                   REGION "TEST STRING TOO LONG"
                       IF LEN(#lengthTest) > #maxLength THEN
                           #_lineBox[#pLineBox] := "Trim"(#_lineBox[#pLineBox]);
                           #_lineBox[#pLineBox] := "Trim"(#_lineBox[#pLineBox]);
                           #pLineBox := #pLineBox + 1;
                           #_lineBox[#pLineBox] := #stringBox[#pString];
                       END_IF;
                   END_REGION

               END_IF;
           END_REGION

       END_FOR;
   END_REGION

   REGION "RETURN"
       #lineBox := #_lineBox;
   END_REGION
END_FUNCTION

FUNCTION "WString.Word_Wrap_Depricated.Concat_Lines" : WString   // FC75, SCL
{ S7_Optimized_Access := 'TRUE' }
VERSION : 0.1
   VAR_INPUT
      lineBox : Array[0..#limitLines] of WString["LONG_STRING_LENGTH"];
   END_VAR
   VAR_TEMP
      pLine : Int;
      ret : WString;
   END_VAR
   VAR CONSTANT
      space : WString := WSTRING#' ';
      blank : WString;
      lineBreak : WString := WSTRING#'$L';
      limitString : Int := 49;
      limitLines : Int := 9;
   END_VAR
BEGIN
   REGION "FOR EACH LINE"
       FOR #pLine := 0 TO #limitLines DO

           REGION "ON END OF LINE LIST"
               IF #lineBox[#pLine] = #space OR #lineBox[#pLine] = #blank THEN
                   EXIT;
               END_IF;
           END_REGION

           REGION "ON FIRST ELEMENT IN LINE LIST"
               IF #pLine = 0 THEN
                   #ret := #lineBox[#pLine];
               END_IF;
           END_REGION

           REGION "CONSTRUCT OUTPUT"
               IF #pLine >= 1 THEN

                   REGION "NO OP ON LINE BREAK CHARACTER"
                       IF #lineBox[#pLine] = #lineBreak THEN
                           ;// no action required
                       END_IF;
                   END_REGION

                   REGION "CONCATINATION"
                       IF #lineBox[#pLine] <> #lineBreak THEN
                           #ret := CONCAT_WSTRING(IN1 := #ret,
                                                  IN2 := #lineBreak,
                                                  IN3 := #lineBox[#pLine]);
                       END_IF;
                   END_REGION

               END_IF;
           END_REGION


       END_FOR;
   END_REGION

   REGION "RETURN"
       #ret := "Trim"(#ret);
       #"WString.Word_Wrap_Depricated.Concat_Lines" := #ret;
   END_REGION
END_FUNCTION

FUNCTION "WString.Split_Single" : Void   // FC202, SCL
{ S7_Optimized_Access := 'TRUE' }
VERSION : 0.1
   VAR_INPUT
      wstring_in : WString;
      delimeter : WString;
      pointer : Int;
   END_VAR
   VAR_IN_OUT
      sub_strings : Array[*] of WString;
   END_VAR
   VAR_TEMP
      _split : WString;
      _position : Int;
      _return : WString;
   END_VAR
BEGIN
   REGION "GET POSITION OF DELIMETER IN STRING"
       #_position := FIND(IN1 := #wstring_in,
                          IN2 := #delimeter);
   END_REGION

   REGION "BASE CASE"
       IF #_position = 0 THEN
           #sub_strings[#pointer] := #wstring_in;
           RETURN;
       END_IF;
   END_REGION


   REGION "RECURSIVE CASE"
       #sub_strings[#pointer] := LEFT(IN := #wstring_in, L := #_position - 1);
       "WString.Split_Single"(wstring_in := RIGHT(IN := #wstring_in, L := LEN(#wstring_in) - #_position),
                       delimeter := #delimeter,
                       "pointer" := #pointer + 1,
                       sub_strings := #sub_strings);
   END_REGION
END_FUNCTION

FUNCTION "WString.Word_Wrap" : WString   // FC203, SCL
{ S7_Optimized_Access := 'TRUE' }
VERSION : 0.1
   VAR_INPUT
      delimeters : Array[*] of WString[1];
      line_length : Int;
      wstring_in : WString;
   END_VAR
   VAR_TEMP
      _i : Int;
      _substring_length : Int;
      _wstring_in_length : Int;
      _pointer_substrings : Int;
      _substring : WString;
      _position_of_last_delimeter : Int;
      _recurse : Bool;
      _string_split_right : WString;
   END_VAR
   VAR CONSTANT
      BLANK : WString;
      NEW_LINE : WString := WSTRING#'$L';
   END_VAR
BEGIN
   #_wstring_in_length := LEN(#wstring_in);

   IF #line_length = 0 THEN
       #"WString.Word_Wrap" := #BLANK;
       RETURN;
   END_IF;

   FOR #_i := 1 TO #_wstring_in_length DO

       #_substring := CONCAT_WSTRING(IN1 := #_substring,
                                     IN2 := #wstring_in[#_i]);
       #_substring_length := LEN(#_substring);

       IF "Array.WString.Is_Element"(search_term := #wstring_in[#_i], search_array := #delimeters) THEN
           #_position_of_last_delimeter := #_i;
       END_IF;

       IF #wstring_in[#_i] = #NEW_LINE THEN
           #_substring := LEFT_WSTRING(IN := #_substring,
                                       L := #_substring_length - 1);
           #_string_split_right := RIGHT_WSTRING(IN := #wstring_in,
                                                 L := #_wstring_in_length - #_i);
           #_recurse := TRUE;
       END_IF;

       IF (#_substring_length = #line_length) AND (#_position_of_last_delimeter <> 0) THEN
           #_substring := LEFT_WSTRING(IN := #_substring,
                                       L := #_position_of_last_delimeter);
           #_string_split_right := RIGHT_WSTRING(IN := #wstring_in,
                                                 L := #_wstring_in_length - #_position_of_last_delimeter);
           #_recurse := TRUE;
       END_IF;

       IF (#_substring_length = #line_length) AND (#_position_of_last_delimeter = 0) THEN
           #_string_split_right := RIGHT_WSTRING(IN := #wstring_in,
                                                 L := #_wstring_in_length - #_substring_length);
           #_recurse := TRUE;
       END_IF;

       IF #_recurse THEN
           #_substring := CONCAT_WSTRING(IN1 := "Trim"(#_substring),
                                         IN2 := #NEW_LINE,
                                         IN3 := "WString.Word_Wrap"(delimeters := #delimeters,
                                                                    line_length := #line_length,
                                                                    wstring_in := #_string_split_right));
           #"WString.Word_Wrap" := #_substring;
           RETURN;
       END_IF;

   END_FOR; 

   #"WString.Word_Wrap" := "Trim"(#_substring);
END_FUNCTION

FUNCTION "WString.Find_Multiple.Depth" : Int   // FC204, SCL
{ S7_Optimized_Access := 'TRUE' }
VERSION : 0.1
   VAR_INPUT
      body : WString;
      terms : Array[*] of WString;
      p_terms : Int;
   END_VAR
   VAR_TEMP
      _length : UDInt;
      _position : Int;
   END_VAR
   VAR CONSTANT
      BLANK : WString;
   END_VAR
BEGIN
   (* 
       Depth first search of 'body' for first occurance of any element of 'terms'.
       For breadth first search, use WString.Find_Multiple.Breadth.
       Returns character postion in the string (1 indexed).
       E.G.: 
           - body := WSTRING#'today?'
           - terms := <WSTRING#>['?', 'ay']
           - returns --> 6
       E.G.:
           - body := WSTRING#'today?'
           - terms := <WSTRING#>['ay', '?']
           - returns --> 4
   *)

   #_length := "Array.Any.Length"(#terms);

   IF #p_terms > #_length OR #terms[#p_terms] = #BLANK THEN
           #"WString.Find_Multiple.Depth" := 0;
       RETURN;
   END_IF;

   #_position := FIND(IN1 := #body,
                      IN2 := #terms[#p_terms]);

   IF #_position = 0 THEN
       #_position := "WString.Find_Multiple.Depth"(body := #body,
                                             terms := #terms,
                                             p_terms := #p_terms + 1);
   END_IF;

   #"WString.Find_Multiple.Depth" := #_position;
END_FUNCTION

FUNCTION "WString.Find_Multiple.Breadth" : Int   // FC205, SCL
{ S7_Optimized_Access := 'TRUE' }
VERSION : 0.1
   VAR_INPUT
      body : WString;
      terms : Array[*] of WString[1];
   END_VAR
   VAR_TEMP
      _i : Int;
      _length : UDInt;
      _min : Int;
      _position : Int;
   END_VAR
   VAR CONSTANT
      BLANK : WString;
   END_VAR
BEGIN
   (* 
       Depth first search of 'body' for first occurance of any element of 'terms'.
       For depth first search use WString.Find_Multiple.Depth.
       Returns character postion in the string (1 indexed).
       E.G.: 
           - body := WSTRING#'today?'
           - terms := <WSTRING#>['?', 'ay']
           - returns --> 6
       E.G.:
           - body := WSTRING#'today?'
           - terms := <WSTRING#>['ay', '?']
           - returns --> 4
   *)

   #_length := "Array.Any.Length"(#terms);

   IF #_length = 0 OR #body = #BLANK THEN
       #"WString.Find_Multiple.Breadth" := 0;
       RETURN;
   END_IF;

   FOR #_i := 0 TO UDINT_TO_INT(#_length) - 1 DO
       #_position := FIND(IN1 := #body,
                          IN2 := #terms[#_i]);
       IF #_position = 0 THEN
           CONTINUE;
       END_IF;
       IF #_position < #_min OR #_min = 0 THEN
           #_min := #_position;
       END_IF;
   END_FOR;

   #"WString.Find_Multiple.Breadth" := #_min;
END_FUNCTION

FUNCTION "WString.Split_Multiple" : Void   // FC206, SCL
{ S7_Optimized_Access := 'TRUE' }
VERSION : 0.1
   VAR_INPUT
      wstring_in : WString;
      delimeters : Array[*] of WString[1];
      pointer : Int;
   END_VAR
   VAR_OUTPUT
      substrings : Array[*] of WString[20];
   END_VAR
   VAR_TEMP
      _i : Int;
      _position : Int;
      _return : WString;
      _split : WString;
   END_VAR
BEGIN
   REGION "GET POSITION OF DELIMETER IN STRING"
       #_position := "WString.Find_Multiple.Breadth"(body := #wstring_in,
                                                     terms := #delimeters);
   END_REGION

   REGION "BASE CASE"
       IF #_position = 0 THEN
           #substrings[#pointer] := #wstring_in;
           "WString.Split_Multiple.Clean_Output"("pointer" := #pointer + 1,
                                                 substrings := #substrings);
           RETURN;
       END_IF;
   END_REGION


   REGION "RECURSIVE CASE"
       #substrings[#pointer] := LEFT(IN := #wstring_in, L := #_position);
       "WString.Split_Multiple"(wstring_in := RIGHT(IN := #wstring_in, L := LEN(#wstring_in) - #_position),
                                delimeters := #delimeters,
                                "pointer" := #pointer + 1,
                                substrings => #substrings);
   END_REGION
END_FUNCTION

FUNCTION "WString.Split_Multiple.Clean_Output" : Void   // FC208, SCL
{ S7_Optimized_Access := 'TRUE' }
VERSION : 0.1
   VAR_INPUT
      pointer : Int;
   END_VAR
   VAR_IN_OUT
      substrings : Array[*] of WString;
   END_VAR
   VAR_TEMP
      _i : Int;
   END_VAR
   VAR CONSTANT
      BLANK : WString;
   END_VAR
BEGIN
   FOR #_i := #"pointer" TO UDINT_TO_INT("Array.Any.Length"(#substrings)) - 1 DO
       #substrings[#_i] := wstring#'';
   END_FOR;
END_FUNCTION

// folder: Utilities/Table Navigation

FUNCTION_BLOCK "Table Nav: End of Data Rollover"   // FB11, SCL
{ S7_Optimized_Access := 'TRUE' }
VERSION : 0.1
   VAR_INPUT
      tblData : Variant;
      tblDisp : Variant;
      nullFlag : Int;
      nullCheck : Variant;
      tableNav : "Nav Bar Data: PLC";
   END_VAR
   VAR_IN_OUT
      rowIndices : Variant;
   END_VAR
   VAR_TEMP
      firstNullIndex : DInt;
      len : Struct
         tblData : DInt;
         tblDisp : DInt;
      END_STRUCT;
      nullCheckVals : Array[0..#lenArrs] of DInt;
      offset : DInt;
      pulses : "Nav Bar Data: PLC";
      RET_VAL : Int;
      retRowIndices : Array[0..#lenArrs] of DInt;
   END_VAR
   VAR CONSTANT
      lenArrs : DInt := 999;
   END_VAR
BEGIN
       REGION "DESCRIPTION"
           (*
           Double checks row indicies against data and rolls over on end of data flag.
           *)
       END_REGION

       REGION "COPY TO LOCAL"
           #RET_VAL := MOVE_BLK_VARIANT(SRC := #rowIndices,
                                        COUNT := CountOfElements(#rowIndices),
                                        SRC_INDEX := 0,
                                        DEST_INDEX := 0,
                                        DEST => #retRowIndices);
           #RET_VAL := MOVE_BLK_VARIANT(SRC := #nullCheck,
                                        COUNT := CountOfElements(#nullCheck),
                                        SRC_INDEX := 0,
                                        DEST_INDEX := 0,
                                        DEST => #nullCheckVals);
       END_REGION

       REGION "GET ARRAY PARAMETERS"
           #len.tblData := UDINT_TO_DINT(CountOfElements(#tblData));
           #len.tblDisp := UDINT_TO_DINT(CountOfElements(#tblDisp));
       END_REGION

       REGION "CALCUALTE ROW INDICIES"
           "Table Nav: Calc Row Indices"(lenTblData := #firstNullIndex,
                                         lenTblDisp := #len.tblDisp,
                                         r1 := #retRowIndices[0],
                                         rowIndicies := #retRowIndices);
       END_REGION

       REGION "RETURN ROW INDICIES"
           #RET_VAL := MOVE_BLK_VARIANT(SRC := #retRowIndices,
                                        COUNT := DINT_TO_UDINT(#len.tblDisp),
                                        SRC_INDEX := 0,
                                        DEST_INDEX := 0,
                                        DEST => #rowIndices);
       END_REGION
END_FUNCTION_BLOCK

FUNCTION_BLOCK "Table Nav"   // FB43, SCL
{ S7_Optimized_Access := 'TRUE' }
VERSION : 0.1
   VAR_INPUT
      first_null_index : DInt;   // if you want to roll over before the end of your array, find the first null index and enter it here
      tblData : Variant;   // array to scan
      tblDisp : Variant;   // viewport array
      tableNav : "Nav Bar Data: PLC";   // table navigation udt
   END_VAR
   VAR_IN_OUT
      rowIndices : Variant;
   END_VAR
   VAR
      "inst Pulses: Table Nav" : "Table Nav: Pulses";
      r1 : DInt;
   END_VAR
   VAR_TEMP
      len : Struct
         tblData : DInt;
         tblDisp : DInt;
      END_STRUCT;
      offset : DInt;
      pulses : "Nav Bar Data: PLC";
      RET_VAL : Int;
      ret_row_indices : Array[0..#lenArrs] of DInt;
      ubound : DInt;
   END_VAR
   VAR CONSTANT
      lenArrs : DInt := 999;
   END_VAR
BEGIN
   REGION "DESCRIPTION"
       (*
       The function returns row indicies indicating the visible rows of a larger
       table determined by standard table navigation buttons.
       The function uses the variant data type to handle tables of any size.
       Rollover and rollunder features are built in.
       Row indices must be output to an array of dint (dimension is flexible).
       *)
   END_REGION


   REGION "GET PRESS PULSES"    
       #"inst Pulses: Table Nav"(press := #tableNav,
                                 pulses => #pulses);
   END_REGION


   REGION "RUN ON BUTTON PRESS"
       IF "Table Nav: Run Trigger"(#pulses) THEN

           REGION "GET ARRAY PARAMETERS"
               #len.tblData := UDINT_TO_DINT(CountOfElements(#tblData));
               #len.tblDisp := UDINT_TO_DINT(CountOfElements(#tblDisp));
           END_REGION

           REGION "CALCULATE UPPER BOUND"
               #ubound := #len.tblData;
               IF #first_null_index <= #len.tblData THEN
                   IF #first_null_index > 0 THEN
                       #ubound := #first_null_index;
                   END_IF;
               END_IF;
           END_REGION


           REGION "CALCULATE OFFSET"
               #offset := "Table Nav: Calculate Offset"(pulses := #pulses,
                                                        lenTblData := #ubound,
                                                        lenTblDisp := #len.tblDisp,
                                                        r1 := #r1);
           END_REGION


           REGION "CALCULATE FIRST ROW"
               #r1 := "Table Nav: Get First Row"(table_length := #ubound,
                                                 offset := #offset,
                                                 first_row := #r1);
           END_REGION


           REGION "CALCUALTE ROW INDICIES"
               "Table Nav: Calc Row Indices"(lenTblData := #ubound,
                                             lenTblDisp := #len.tblDisp,
                                             r1 := #r1,
                                             rowIndicies := #ret_row_indices);
           END_REGION


           REGION "RETURN ROW INDICIES"
               #RET_VAL := MOVE_BLK_VARIANT(SRC := #ret_row_indices,
                                            COUNT := DINT_TO_UDINT(#len.tblDisp),
                                            SRC_INDEX := 0,
                                            DEST_INDEX := 0,
                                            DEST => #rowIndices);
           END_REGION

       END_IF;
   END_REGION
END_FUNCTION_BLOCK

FUNCTION_BLOCK "Table Nav: Pulses"   // FB44, SCL
{ S7_Optimized_Access := 'TRUE' }
VERSION : 0.1
   VAR_INPUT
      press : "Nav Bar Data: PLC";
   END_VAR
   VAR_OUTPUT
      pulses : "Nav Bar Data: PLC";
   END_VAR
   VAR
      old : "Nav Bar Data: PLC";
   END_VAR
BEGIN
   REGION "EVALUATION"
       #pulses.top.actuate := #press.top.actuate AND NOT #old.top.actuate;
       #pulses.pageUp.actuate := #press.pageUp.actuate AND NOT #old.pageUp.actuate;
       #pulses.lineUp.actuate := #press.lineUp.actuate AND NOT #old.lineUp.actuate;
       #pulses.lineDown.actuate := #press.lineDown.actuate AND NOT #old.lineDown.actuate;
       #pulses.pageDown.actuate := #press.pageDown.actuate AND NOT #old.pageDown.actuate;
       #pulses.bottom.actuate := #press.bottom.actuate AND NOT #old.bottom.actuate;
   END_REGION

   REGION "CHANGE DETECTION"
       #old.top.actuate := #press.top.actuate;
       #old.pageUp.actuate := #press.pageUp.actuate;
       #old.lineUp.actuate := #press.lineUp.actuate;
       #old.lineDown.actuate := #press.lineDown.actuate;
       #old.pageDown.actuate := #press.pageDown.actuate;
       #old.bottom.actuate := #press.bottom.actuate;
   END_REGION
END_FUNCTION_BLOCK

FUNCTION "Table Nav: Get Null Index" : DInt   // FC14, SCL
{ S7_Optimized_Access := 'TRUE' }
VERSION : 0.1
   VAR_INPUT
      nullFlag : Int;
      nullCheckVals : Array[0.."WIP_COUNT"] of DInt;
   END_VAR
   VAR_TEMP
      pNullCheck : DInt;
   END_VAR
BEGIN
   WHILE #nullCheckVals[#pNullCheck] <> #nullFlag AND #pNullCheck <= "WIP_COUNT" DO
       #pNullCheck += 1;
   END_WHILE;
   #"Table Nav: Get Null Index" := #pNullCheck;
END_FUNCTION

FUNCTION "Table Nav: Get First Row" : DInt   // FC44, SCL
{ S7_Optimized_Access := 'TRUE' }
VERSION : 0.1
   VAR_INPUT
      first_row : DInt;
      offset : DInt;
      table_length : DInt;
   END_VAR
   VAR_TEMP
      ret : DInt;
   END_VAR
BEGIN
   REGION "DESCRIPTION"
       (*
       The new first row of the table is calculated from the offset. 
       Rollover and rollunder are resolved for the first row.
       *)
   END_REGION

   REGION "COPY TO INTERNAL"
       #ret := #first_row + #offset;
   END_REGION

   REGION "ROLLUNDER"
       IF #ret < 0 THEN
           #ret := #ret + #table_length;
       END_IF;
   END_REGION

   REGION "ROLLOVER"
       IF #ret > #table_length THEN
           #ret := #ret - #table_length;
       END_IF;
   END_REGION

   REGION "OUTPUT"
       #"Table Nav: Get First Row" := #ret;
   END_REGION
END_FUNCTION

FUNCTION "Table Nav: Calculate Offset" : DInt   // FC45, SCL
{ S7_Optimized_Access := 'TRUE' }
VERSION : 0.1
   VAR_INPUT
      lenTblData : DInt;
      lenTblDisp : DInt;
      pulses : "Nav Bar Data: PLC";
      r1 : DInt;
   END_VAR
   VAR_TEMP
      retOffset : DInt;
   END_VAR
   // Ret_Val : offset from table row 1 from button
BEGIN
   REGION "DESCRIPTION"
       (*
       The offset from the first row of the table is calculated based on the button pressed.
       *)
   END_REGION

   REGION "TOP"
       IF #pulses.top.actuate THEN
           #retOffset := -1 * #r1;
       END_IF;
   END_REGION

   REGION "PAGE UP"
       IF #pulses.pageUp.actuate THEN
           #retOffset := -1 * #lenTblDisp;
       END_IF;
   END_REGION

   REGION "LINE UP"
       IF #pulses.lineUp.actuate THEN
           #retOffset := -1;
       END_IF;
   END_REGION

   REGION "LINE DOWN"
       IF #pulses.lineDown.actuate THEN
           #retOffset := 1;
       END_IF;
   END_REGION

   REGION "PAGE DOWN"
       IF #pulses.pageDown.actuate THEN
           #retOffset := #lenTblDisp ;
       END_IF;
   END_REGION

   REGION "BOTTOM"
       IF #pulses.bottom.actuate THEN
           #retOffset := #lenTblData - #lenTblDisp - #r1;
       END_IF;
   END_REGION

   REGION "RETURN"
       #"Table Nav: Calculate Offset" := #retOffset;
   END_REGION
END_FUNCTION

FUNCTION "Table Nav: Calc Row Indices" : Void   // FC46, SCL
{ S7_Optimized_Access := 'TRUE' }
VERSION : 0.1
   VAR_INPUT
      lenTblData : DInt;
      lenTblDisp : DInt;
      r1 : DInt;
   END_VAR
   VAR_IN_OUT
      rowIndicies : Array[0..#lenRetArr] of DInt;
   END_VAR
   VAR_TEMP
      pOutArr : Int;
      calcRowIdx : DInt;
      retRowIndicies : Array[0..#lenRetArr] of DInt;
   END_VAR
   VAR CONSTANT
      lenRetArr : Int := 999;
   END_VAR
BEGIN
   REGION "DESCRIPTION"
       (*
       An array of the row indicies that the table should display is returned.
       Rollover and rollunder are calculated index by index.
       *) 
   END_REGION

   REGION "INITIALIZE OUTPUT"
       FOR #pOutArr := 0 TO #lenRetArr DO
           #rowIndicies[#pOutArr] := 0;
       END_FOR;
   END_REGION

   REGION "CALCULATE INDICIES"
       FOR #pOutArr := 0 TO DINT_TO_INT(#lenTblDisp) DO

           REGION "CALCULATE INDEX"
               #calcRowIdx := #r1 + INT_TO_DINT(#pOutArr);
           END_REGION

           REGION "ROLL UNDER"
               IF #calcRowIdx < 0 THEN
                   #calcRowIdx := #calcRowIdx + #lenTblDisp;
               END_IF;
           END_REGION

           REGION "ROLL OVER"
               IF #calcRowIdx >= #lenTblData THEN
                   #calcRowIdx := #calcRowIdx - #lenTblData;
               END_IF;
           END_REGION

           REGION "SAVE TO ARRAY"
               #retRowIndicies[#pOutArr] := #calcRowIdx;
           END_REGION

       END_FOR;
   END_REGION

   REGION "OUTPUT"
       #rowIndicies := #retRowIndicies;
   END_REGION
END_FUNCTION

FUNCTION "Table Nav: Run Trigger" : Bool   // FC47, SCL
{ S7_Optimized_Access := 'TRUE' }
VERSION : 0.1
   VAR_INPUT
      pulses : "Nav Bar Data: PLC";
   END_VAR
BEGIN
   #"Table Nav: Run Trigger" :=
       #pulses.top.actuate OR
       #pulses.pageUp.actuate OR
       #pulses.lineUp.actuate OR
       #pulses.lineDown.actuate OR
       #pulses.pageDown.actuate OR
       #pulses.bottom.actuate;
END_FUNCTION

// folder: Utilities/Timer

FUNCTION "Timer.Time_to_WString" : WString   // FC36, SCL
{ S7_Optimized_Access := 'TRUE' }
VERSION : 0.1
   VAR_INPUT
      "Time" : Time;
   END_VAR
   VAR_TEMP
      "Time as DInt" : DInt;
      "Hours 10s Place" : DInt;
      "Hours 1s Place" : DInt;
      "Minutes 10s Place" : DInt;
      "Minutes 1s Place" : DInt;
      "Seconds 10s Place" : DInt;
      "Seconds 1s Place" : DInt;
      "Time Elements" : Array[0..4] of WString;
      Length : Int;
      "String Box" : WString;
      "DInt Box" : DInt;
   END_VAR
   VAR CONSTANT
      "Milliseconds per 10 Hours" : DInt := 36_000_000;
      "Milliseconds per Hour" : DInt := 3_600_000;
      "Milliseconds per 10 Minutes" : DInt := 600_000;
      "Milliseconds per Minute" : DInt := 60_000;
      "Milliseconds per 10 Seconds" : DInt := 10_000;
      "Milliseconds per Second" : DInt := 1_000;
   END_VAR
BEGIN
   REGION GET INPUT
       #"Time as DInt" := #Time;
   END_REGION

   REGION CONVERT TIME INTO INDIVIDUAL PLACE VALUES
       #"Minutes 10s Place" := #"Time as DInt" / #"Milliseconds per 10 Minutes";
       #"Minutes 1s Place" := (#"Time as DInt" / #"Milliseconds per Minute") MOD 10;
       #"Seconds 10s Place" := (#"Time as DInt" MOD #"Milliseconds per Minute") / #"Milliseconds per 10 Seconds";
       #"Seconds 1s Place" := (#"Time as DInt" / #"Milliseconds per Second") MOD 10;
   END_REGION

   REGION "ADD SIGN"
       #"Time Elements"[0] := wstring#'';
       IF #"Minutes 10s Place" < 0 OR
           #"Minutes 1s Place" < 0 OR
           #"Seconds 10s Place" < 0 OR
           #"Seconds 1s Place" < 0 THEN
            #"Time Elements"[0] := wstring#'-';
       END_IF;
   END_REGION

   REGION CONVERT PLACE VALUES INTO COMPONENT STRINGS
       // MINUTES
       #"DInt Box" := #"Minutes 10s Place" * 10 + #"Minutes 1s Place";
       #"String Box" := DINT_TO_WSTRING(IN := #"DInt Box");
       #"String Box" := "Strip Sign"("WString":=#"String Box");
       #"String Box" := "Add Leading"("Leading Character" := WCHAR#'0',
                                      "Desired Length" := 2,
                                      "String" := #"String Box");
       #"Time Elements"[1] := #"String Box";
       // COLON
       #"Time Elements"[2] := WSTRING#':';
       // SECONDS
       #"DInt Box" := #"Seconds 10s Place" * 10 + #"Seconds 1s Place";
       #"String Box" := DINT_TO_WSTRING(IN := #"DInt Box");
       #"String Box" := "Strip Sign"("WString":=#"String Box");
       #"String Box" := "Add Leading"("Leading Character" := WCHAR#'0',
                                      "Desired Length" := 2,
                                      "String" := #"String Box");
       #"Time Elements"[3] := #"String Box";
   END_REGION


   REGION RETURN VALUE
       #"Timer.Time_to_WString" := CONCAT_WSTRING(IN1 := #"Time Elements"[0],
                                            IN2 := #"Time Elements"[1],
                                            IN3 := #"Time Elements"[2],
                                            IN4 := #"Time Elements"[3]);
   END_REGION
END_FUNCTION

FUNCTION "Timer.WString_to_Time" : Time   // FC38, SCL
{ S7_Optimized_Access := 'TRUE' }
VERSION : 0.1
   VAR_INPUT
      WString : WString;
   END_VAR
   VAR_TEMP
      Count : UInt;
      "DInt Box" : DInt;
      "String Box" : WString [5];
      "Time Box" : Time;
      "WChar Array" : Array[0..4] of WChar;
   END_VAR
   VAR CONSTANT
      "ms/(10 hr)" : DInt := 36_000_000;
      "ms/hr" : DInt := 3_600_000;
      "ms/(10 min)" : DInt := 600_000;
      "ms/min" : DInt := 60_000;
      "ms/(10 sec)" : DInt := 10_000;
      "ms/sec" : DInt := 1_000;
   END_VAR
BEGIN
   REGION EXPLODE INPUT

       #"String Box" := #WString;
       IF #"String Box" = WSTRING#'' THEN
           #"String Box" := WSTRING#'00:00';
       END_IF;

       Strg_TO_Chars(Strg := #"String Box",
                     pChars := 0,
                     Cnt => #Count,
                     Chars := #"WChar Array");

   END_REGION

   REGION CONVERT ARRAY ELEMENTS TO TIME

       // 10S OF MINUTES
       #"DInt Box" := WCHAR_TO_DINT(IN := #"WChar Array"[0]) - 16#30;
       #"Time Box" := #"Time Box" + #"DInt Box" * #"ms/(10 min)";

       // MINUTES
       #"DInt Box" := WCHAR_TO_DINT(IN := #"WChar Array"[1]) - 16#30;
       #"Time Box" := #"Time Box" + #"DInt Box" * #"ms/min";

       // 10S OF SECONDS
       #"DInt Box" := WCHAR_TO_DINT(IN := #"WChar Array"[3]) - 16#30;
       #"Time Box" := #"Time Box" + #"DInt Box" * #"ms/(10 sec)";

       // SECONDS
       #"DInt Box" := WCHAR_TO_DINT(IN := #"WChar Array"[4]) - 16#30;
       #"Time Box" := #"Time Box" + #"DInt Box" * #"ms/sec";

   END_REGION


   REGION RETURN VALUE

       #"Timer.WString_to_Time" := #"Time Box";

   END_REGION
END_FUNCTION

FUNCTION "Timer.WString_to_Real" : Real   // FC39, SCL
{ S7_Optimized_Access := 'TRUE' }
VERSION : 0.1
   VAR_INPUT
      wstring : WString;
   END_VAR
   VAR CONSTANT
      msPerSec : Real := 1000.0;
   END_VAR
BEGIN
   #"Timer.WString_to_Real" := DINT_TO_REAL(TIME_TO_DINT("Timer.WString_to_Time"(#wstring))) / #msPerSec;
END_FUNCTION

FUNCTION "Timer.Real_to_WString" : WString   // FC40, SCL
{ S7_Optimized_Access := 'TRUE' }
VERSION : 0.1
   VAR_INPUT
      realVal : Real;
   END_VAR
   VAR CONSTANT
      msPerSec : Real := 1000.0;
   END_VAR
BEGIN
   #"Timer.Real_to_WString" := "Timer.Time_to_WString"(DINT_TO_TIME(REAL_TO_DINT(#realVal * #msPerSec)));
END_FUNCTION

FUNCTION "Timer" : Void   // FC79, SCL
{ S7_Optimized_Access := 'TRUE' }
VERSION : 0.1
   VAR_INPUT
      delta : Real;
      allotted : Real;
   END_VAR
   VAR_IN_OUT
      elapsed : Real;
      remaining : Real;
   END_VAR
   VAR_TEMP
      _elapsed : Real;
      _remaining : Real;
   END_VAR
BEGIN
   #_elapsed := #elapsed + #delta;
   #_remaining := #allotted - #_elapsed;
   #elapsed := #_elapsed;
   #remaining := #_remaining;
END_FUNCTION

// folder: Utilities/UInt

FUNCTION "UInt.Value_Change" : Bool   // FC183, SCL
{ S7_Optimized_Access := 'TRUE' }
VERSION : 0.1
   VAR_INPUT
      value : UInt;
      old_value : UInt;
   END_VAR
BEGIN
   #"UInt.Value_Change" := #value <> #old_value;
END_FUNCTION

// folder: Utilities/WIP

FUNCTION "WIP.Code_to_WString" : WString   // FC64, SCL
{ S7_Optimized_Access := 'TRUE' }
VERSION : 0.1
   VAR_INPUT
      wipTxtLib : "Recipe: Wip Text Library";
      code : DInt;
   END_VAR
   VAR_TEMP
      wipCode : DInt;
      wipText : DInt;
      output : WString;
   END_VAR
   VAR CONSTANT
      newLine : WString := WSTRING#'$L';
   END_VAR
BEGIN
   REGION "PARSE CODE"
       "Part_Number.Parse_Code"(code := #code,
                    code_left => #wipCode,
                    code_right => #wipText);
   END_REGION

   REGION "DOUBLE LINE PN"
       #output := CONCAT_WSTRING(IN1 := #wipTxtLib.code[#wipCode],
                                 IN2 := #newLine,
                                 IN3 := #wipTxtLib.txt[#wipText]);
   END_REGION

   REGION "OUTPUT"
       #"WIP.Code_to_WString" := #output;
   END_REGION
END_FUNCTION

FUNCTION "WIP.Count" : Int   // FC72, SCL
{ S7_Optimized_Access := 'TRUE' }
VERSION : 0.1
   VAR_INPUT
      stnSavedWips : "WIP: Station";
   END_VAR
   VAR_TEMP
      pWip : Int;
   END_VAR
   // Ret_Val : -1 for no wips in station
BEGIN
   WHILE #stnSavedWips.wip[#pWip].wip.code <> -1 DO
       #pWip += 1;
   END_WHILE;
   #"WIP.Count" := #pWip - 1;
END_FUNCTION

FUNCTION "WIP.Global_Index_to_Station" : "WIP: Station"   // FC113, SCL
{ S7_Optimized_Access := 'TRUE' }
VERSION : 0.1
   VAR_INPUT
      index : Int;
      wip_stations : "Recipe: HMI Stations Saved Wips";
   END_VAR
   VAR_TEMP
      i : Int;
      ret : "WIP: Station";
   END_VAR
BEGIN
   REGION "FIND STATION"
       FOR #i := 0 TO "HMI_STATION_COUNT" DO
           IF #wip_stations.stn[#i].pStn = #index THEN
               #ret := #wip_stations.stn[#i];
               EXIT;
           END_IF;
       END_FOR;
   END_REGION


   REGION "RETURN"
       #"WIP.Global_Index_to_Station" := #ret;
   END_REGION
END_FUNCTION

FUNCTION "WIP.Global_Index_to_HMI_Station_Index" : Int   // FC130, SCL
{ S7_Optimized_Access := 'TRUE' }
VERSION : 0.1
   VAR_INPUT
      global_index : Int;
      saved_WIPs : "Recipe: HMI Stations Saved Wips";
   END_VAR
   VAR_TEMP
      i : Int;
      ret : Int;
   END_VAR
BEGIN
   REGION "SEARCH FOR INDEX"
       #ret := "NULL_TOKEN";
       FOR #i := 0 TO "HMI_STATION_COUNT" DO
           IF #saved_WIPs.stn[#i].pStn = #global_index THEN
               #ret := #i;
               EXIT;
           END_IF;
       END_FOR;
   END_REGION


   REGION "RETURN"
       #"WIP.Global_Index_to_HMI_Station_Index" := #ret;
   END_REGION
END_FUNCTION

FUNCTION "WIP.Code_to_Index" : Int   // FC233, SCL
{ S7_Optimized_Access := 'TRUE' }
VERSION : 0.1
   VAR_INPUT
      saved_wip : "WIP: Station";
      wip_code : DInt;
   END_VAR
   VAR_TEMP
      _i : Int;
      _length : Int;
   END_VAR
BEGIN
   #_length := UDINT_TO_INT("Array.Any.Length"(#saved_wip.wip)) - 1;
   FOR #_i := 0 TO #_length DO
       IF #wip_code <> #saved_wip.wip[#_i].wip.code THEN
           CONTINUE;
       END_IF;
       #"WIP.Code_to_Index" := #_i;
       RETURN;
   END_FOR;

   #"WIP.Code_to_Index" := "NULL_TOKEN";
   RETURN;
END_FUNCTION

FUNCTION "WIP_Station.Indices_of_Selected_WIPs" : Void   // FC241, SCL
{ S7_Optimized_Access := 'TRUE' }
VERSION : 0.1
   VAR_INPUT
      selected_wips : "Selected Wips";
      station_wips : "WIP: Station";
   END_VAR
   VAR_IN_OUT
      selected_wip_indices : Array[*] of Int;
   END_VAR
   VAR_TEMP
      _i : Int;
      _length : Int;
      _p_return : Int;
      _wip_index : Int;
   END_VAR
   VAR CONSTANT
      UBOUND : Int := 999;
   END_VAR
BEGIN
   REGION "PREP ARRAY OF FOUND INDICES"
       "Array.Int.Fill"(value := "NULL_TOKEN",
                        int_array := #selected_wip_indices);
       #_length := UDINT_TO_INT("Array.Any.Length"(#selected_wip_indices)) - 1;
   END_REGION

   REGION "FOR EACH SELECTED WIP"
       FOR #_i := 0 TO #selected_wips.count - 1 DO

           REGION "GET SELECTED WIPS INDEX IN THIS STATION"
               #_wip_index := "WIP_Station.Indices_of_Selected_WIPS.Search_WIP"(wip_code := #selected_wips.wips[#_i],
                                                                                station_wips := #station_wips);
           END_REGION

           REGION "IF NOT FOUND GO TO NEXT WIP"
               // fault tolerance
               IF #_wip_index = "NULL_TOKEN" THEN
                   CONTINUE;
               END_IF;
           END_REGION

           REGION "WIP FOUND IN STATION"
               #selected_wip_indices[#_p_return] := #_wip_index;
               #_p_return += 1;
           END_REGION

           REGION "DON'T GO OUT OF FOUND IDEX ARRAY"
               // fault tolerance
               IF #_p_return > #_length THEN
                   RETURN;
               END_IF;
           END_REGION

       END_FOR;
   END_REGION
END_FUNCTION

FUNCTION "WIP_Station.Indices_of_Selected_WIPS.Search_WIP" : Int   // FC242, SCL
{ S7_Optimized_Access := 'TRUE' }
VERSION : 0.1
   VAR_INPUT
      wip_code : DInt;
      station_wips : "WIP: Station";
   END_VAR
   VAR_TEMP
      _i : Int;
      _length : Int;
   END_VAR
BEGIN
   REGION "FOR EACH WIP IN STATION"
       #_length := UDINT_TO_INT("Array.Any.Length"(#station_wips.wip)) - 1;
       FOR #_i := 0 TO #_length DO

           REGION "WIP CODE DOES NOT MATCH"
               IF #wip_code <> #station_wips.wip[#_i].wip.code THEN
                   CONTINUE;
               END_IF;
           END_REGION

           REGION "WIP CODE MATCHES"
               #"WIP_Station.Indices_of_Selected_WIPS.Search_WIP" := #_i;
               RETURN;
           END_REGION

       END_FOR;
   END_REGION

   REGION "NO MATCH FOUND"
       #"WIP_Station.Indices_of_Selected_WIPS.Search_WIP" := "NULL_TOKEN";
       RETURN;
   END_REGION
END_FUNCTION

// folder: Utilities/WString

FUNCTION "WString: Rising Edge" : Bool   // FC182, SCL
{ S7_Optimized_Access := 'TRUE' }
VERSION : 0.1
   VAR_INPUT
      value : WString;
      old_value : WString;
   END_VAR
   VAR CONSTANT
      blank : WString;
   END_VAR
BEGIN
   #"WString: Rising Edge" := #value <> #blank AND #old_value = #blank;
END_FUNCTION

FUNCTION "WString: Falling Edge" : Bool   // FC188, SCL
{ S7_Optimized_Access := 'TRUE' }
VERSION : 0.1
   VAR_INPUT
      value : WString;
      old_value : WString;
   END_VAR
   VAR CONSTANT
      blank : WString;
   END_VAR
BEGIN
   #"WString: Falling Edge" := #value = #blank AND #old_value <> #blank;
END_FUNCTION

// ===== library types =====

TYPE "PB Data"
   STRUCT
      actuate : Bool;
      animate : USInt;
      enable : Bool;
      label : WString[80];
      listSelect : UInt;
      visible : Bool;
   END_STRUCT;
END_TYPE

TYPE "PB Data: Text Label"
   STRUCT
      actuate : Bool;
      animate : USInt;
      label : WString[20];
   END_STRUCT;
END_TYPE

TYPE "Station Assignment: Button Details Data"
   STRUCT
      alloted : Struct
         animate : USInt;
         value : WString[10];
      END_STRUCT;
      critical : Struct
         animate : USInt;
         value : WString[10];
      END_STRUCT;
      label : Struct
         animate : USInt;
         value : WString[2];
      END_STRUCT;
      partNumber : Struct
         animate : USInt;
         value : WString[40];
      END_STRUCT;
      select : Struct
         actuate : Bool;
         animate : USInt;
      END_STRUCT;
   END_STRUCT;
END_TYPE

TYPE "IO Field Data: Timers"
   STRUCT
      animate : USInt;
      inputFinished : Bool;
      value : WString[5];
   END_STRUCT;
END_TYPE

TYPE "Line Label Data"
   STRUCT
      animate : Struct
         bg : USInt;
         ioField : USInt;
      END_STRUCT;
      inputFinished : Bool;
      value : WString[10];
   END_STRUCT;
END_TYPE

TYPE "Drop Zone Data"
   STRUCT
      animate : Struct
         bg : USInt;
         ioField : USInt;
      END_STRUCT;
      inputFinished : Bool;
      value : WString[10];
   END_STRUCT;
END_TYPE

TYPE "Station Sim Data"
   STRUCT
      stn : Struct
         animate : USInt;
         label : WString[20];
      END_STRUCT;
      btn : Struct
         actuate : Byte;
         animate : Array[0..7] of USInt;
         labels : Array[0..7] of WString [4];
      END_STRUCT;
   END_STRUCT;
END_TYPE

// folder: Main HMI

TYPE "Table Row Data"
   STRUCT
      address : DInt := -1;
      ordered : Bool;
      pbSelection : Struct
         actuate : Bool;
         animate : USInt;
      END_STRUCT;
      rtBackground : Struct
         animate : USInt;
      END_STRUCT;
      tfDropZone : Struct
         animate : USInt;
         value : WString[20];
      END_STRUCT;
      tfLine : Struct
         animate : USInt;
         value : WString[20];
      END_STRUCT;
      tfPartNumber : Struct
         animateDL : USInt;
         animateSL : USInt;
         value : WString[40];
      END_STRUCT;
      tfTime : Struct
         animate : USInt;
         value : WString[20];
      END_STRUCT;
   END_STRUCT;
END_TYPE

(* ===== HMI "HMI_RT_1" =====
system functions are stored by id; their names below are inferred from use
connection "Main HMI": ETHERNET, S7_1500_OMS

HMI tags "Default tag table"
   "Clock_Byte" : Byte = PLC Clock_Byte AT %MB0, 100 ms
   "HMI Data: Warehouse HMI_screenNumber" : Int = PLC "HMI Data: Warehouse HMI".screenNumber AT %DB1.DBW0, 100 ms
   "HMI Data: Warehouse HMI_barcode" : Barcode Screen = PLC "HMI Data: Warehouse HMI".barcode AT %DB1.DBW0, 100 ms
   "HMI Data: Warehouse HMI_tableNav_top" : Push Button Data = PLC "HMI Data: Warehouse HMI".tableNav.top, 100 ms
   "HMI Data: Warehouse HMI_tableNav_pageUp" : Push Button Data = PLC "HMI Data: Warehouse HMI".tableNav.pageUp, 100 ms
   "HMI Data: Warehouse HMI_tableNav_lineUp" : Push Button Data = PLC "HMI Data: Warehouse HMI".tableNav.lineUp, 100 ms
   "HMI Data: Warehouse HMI_tableNav_lineDown" : Push Button Data = PLC "HMI Data: Warehouse HMI".tableNav.lineDown, 100 ms
   "HMI Data: Warehouse HMI_tableNav_pageDown" : Push Button Data = PLC "HMI Data: Warehouse HMI".tableNav.pageDown, 100 ms
   "HMI Data: Warehouse HMI_tableNav_bottom" : Push Button Data = PLC "HMI Data: Warehouse HMI".tableNav.bottom, 100 ms
   "HMI Data: Warehouse HMI_networkHealth_pnioDevices{1}" : Push Button Data = PLC "HMI Data: Warehouse HMI".networkHealth.pnioDevices[1], 100 ms
   "HMI Data: Warehouse HMI_networkHealth_pnioDevices{2}" : Push Button Data = PLC "HMI Data: Warehouse HMI".networkHealth.pnioDevices[2], 100 ms
   "HMI Data: Warehouse HMI_networkHealth_pnioDevices{3}" : Push Button Data = PLC "HMI Data: Warehouse HMI".networkHealth.pnioDevices[3], 100 ms
   "HMI Data: Warehouse HMI_networkHealth_pnioDevices{4}" : Push Button Data = PLC "HMI Data: Warehouse HMI".networkHealth.pnioDevices[4], 100 ms
   "HMI Data: Warehouse HMI_networkHealth_pnioDevices{5}" : Push Button Data = PLC "HMI Data: Warehouse HMI".networkHealth.pnioDevices[5], 100 ms
   "HMI Data: Warehouse HMI_networkHealth_pnioDevices{6}" : Push Button Data = PLC "HMI Data: Warehouse HMI".networkHealth.pnioDevices[6], 100 ms
   "HMI Data: Warehouse HMI_networkHealth_pnioDevices{7}" : Push Button Data = PLC "HMI Data: Warehouse HMI".networkHealth.pnioDevices[7], 100 ms
   "HMI Data: Warehouse HMI_networkHealth_pnioDevices{8}" : Push Button Data = PLC "HMI Data: Warehouse HMI".networkHealth.pnioDevices[8], 100 ms
   "HMI Data: Warehouse HMI_networkHealth_pnioDevices{9}" : Push Button Data = PLC "HMI Data: Warehouse HMI".settings.selectStation, 100 ms
   "HMI Data: Warehouse HMI_networkHealth_pnioDevices{10}" : Push Button Data = PLC "HMI Data: Warehouse HMI".networkHealth.pnioDevices[10], 100 ms
   "HMI Data: Warehouse HMI_networkHealth_pnioDevices{11}" : Push Button Data = PLC "HMI Data: Warehouse HMI".networkHealth.pnioDevices[11], 100 ms
   "HMI Data: Warehouse HMI_networkHealth_pnioDevices{12}" : Push Button Data = PLC "HMI Data: Warehouse HMI".networkHealth.pnioDevices[12], 100 ms
   "HMI Data: Warehouse HMI_networkHealth_pnioDevices{13}" : Push Button Data = PLC "HMI Data: Warehouse HMI".networkHealth.pnioDevices[13], 100 ms
   "HMI Data: Warehouse HMI_networkHealth_pnioDevices{16}" : Push Button Data = PLC "HMI Data: Warehouse HMI".networkHealth.pnioDevices[16], 100 ms
   "HMI Data: Warehouse HMI_networkHealth_pnioDevices{14}" : Push Button Data = PLC "HMI Data: Warehouse HMI".networkHealth.pnioDevices[14], 100 ms
   "HMI Data: Warehouse HMI_networkHealth_pnioDevices{15}" : Push Button Data = PLC "HMI Data: Warehouse HMI".networkHealth.pnioDevices[15], 100 ms
   "HMI Data: Warehouse HMI_networkHealth_pnioDevices{17}" : Push Button Data = PLC "HMI Data: Warehouse HMI".networkHealth.pnioDevices[17], 100 ms
   "HMI Data: Warehouse HMI_networkHealth_pnioDevices{18}" : Push Button Data = PLC "HMI Data: Warehouse HMI".networkHealth.pnioDevices[18], 100 ms
   "HMI Data: Warehouse HMI_networkHealth_pnioDevices{19}" : Push Button Data = PLC "HMI Data: Warehouse HMI".networkHealth.pnioDevices[19], 100 ms
   "HMI Data: Warehouse HMI_networkHealth_pnioDevices{20}" : Push Button Data = PLC "HMI Data: Warehouse HMI".networkHealth.pnioDevices[20], 100 ms
   "HMI Data: Warehouse HMI_networkHealth_pnioDevices{21}" : Push Button Data = PLC "HMI Data: Warehouse HMI".networkHealth.pnioDevices[21], 100 ms
   "HMI Data: Warehouse HMI_networkHealth_pnioDevices{22}" : Push Button Data = PLC "HMI Data: Warehouse HMI".networkHealth.pnioDevices[22], 100 ms
   "HMI Data: Warehouse HMI_networkHealth_pnioDevices{31}" : Push Button Data = PLC "HMI Data: Warehouse HMI".networkHealth.pnioDevices[31], 100 ms
   "HMI Data: Warehouse HMI_networkHealth_pnioDevices{32}" : Push Button Data = PLC "HMI Data: Warehouse HMI".networkHealth.pnioDevices[32], 100 ms
   "HMI Data: Warehouse HMI_networkHealth_pnioDevices{29}" : Push Button Data = PLC "HMI Data: Warehouse HMI".networkHealth.pnioDevices[29], 100 ms
   "HMI Data: Warehouse HMI_networkHealth_pnioDevices{30}" : Push Button Data = PLC "HMI Data: Warehouse HMI".networkHealth.pnioDevices[30], 100 ms
   "HMI Data: Warehouse HMI_networkHealth_pnioDevices{27}" : Push Button Data = PLC "HMI Data: Warehouse HMI".networkHealth.pnioDevices[27], 100 ms
   "HMI Data: Warehouse HMI_networkHealth_pnioDevices{28}" : Push Button Data = PLC "HMI Data: Warehouse HMI".networkHealth.pnioDevices[28], 100 ms
   "HMI Data: Warehouse HMI_networkHealth_pnioDevices{23}" : Push Button Data = PLC "HMI Data: Warehouse HMI".networkHealth.pnioDevices[23], 100 ms
   "HMI Data: Warehouse HMI_networkHealth_pnioDevices{24}" : Push Button Data = PLC "HMI Data: Warehouse HMI".networkHealth.pnioDevices[24], 100 ms
   "HMI Data: Warehouse HMI_networkHealth_pnioDevices{25}" : Push Button Data = PLC "HMI Data: Warehouse HMI".networkHealth.pnioDevices[25], 100 ms
   "HMI Data: Warehouse HMI_networkHealth_pnioDevices{26}" : Push Button Data = PLC "HMI Data: Warehouse HMI".networkHealth.pnioDevices[26], 100 ms
   "HMI Data: Warehouse HMI_networkHealth_pnioDevices{33}" : Push Button Data = PLC "HMI Data: Warehouse HMI".networkHealth.pnioDevices[33], 100 ms
   "HMI Data: Warehouse HMI_networkHealth_pnioDevices{34}" : Push Button Data = PLC "HMI Data: Warehouse HMI".networkHealth.pnioDevices[34], 100 ms
   "HMI Data: Warehouse HMI_networkHealth_pnioDevices{35}" : Push Button Data = PLC "HMI Data: Warehouse HMI".networkHealth.pnioDevices[35], 100 ms
   "HMI Data: Warehouse HMI_networkHealth_pnioDevices{36}" : Push Button Data = PLC "HMI Data: Warehouse HMI".networkHealth.pnioDevices[36], 100 ms
   "HMI Data: Warehouse HMI_networkHealth_pnioDevices{37}" : Push Button Data = PLC "HMI Data: Warehouse HMI".networkHealth.pnioDevices[37], 100 ms
   "HMI Data: Warehouse HMI_networkHealth_pnioDevices{38}" : Push Button Data = PLC "HMI Data: Warehouse HMI".networkHealth.pnioDevices[38], 100 ms
   "HMI Data: Warehouse HMI_networkHealth_pnioDevices{39}" : Push Button Data = PLC "HMI Data: Warehouse HMI".networkHealth.pnioDevices[39], 100 ms
   "HMI Data: Warehouse HMI_networkHealth_pnioDevices{40}" : Push Button Data = PLC "HMI Data: Warehouse HMI".networkHealth.pnioDevices[40], 100 ms
   "HMI Data: Warehouse HMI_networkHealth_pnioDevices{41}" : Push Button Data = PLC "HMI Data: Warehouse HMI".networkHealth.pnioDevices[41], 100 ms
   "HMI Data: Warehouse HMI_networkHealth_pnioDevices{42}" : Push Button Data = PLC "HMI Data: Warehouse HMI".networkHealth.pnioDevices[42], 100 ms
   "HMI Data: Warehouse HMI_networkHealth_pnioDevices{43}" : Push Button Data = PLC "HMI Data: Warehouse HMI".networkHealth.pnioDevices[43], 100 ms
   "HMI Data: Warehouse HMI_networkHealth_pnioDevices{44}" : Push Button Data = PLC "HMI Data: Warehouse HMI".networkHealth.pnioDevices[44], 100 ms
   "HMI Data: Warehouse HMI_networkHealth_pnioDevices{45}" : Push Button Data = PLC "HMI Data: Warehouse HMI".networkHealth.pnioDevices[45], 100 ms
   "HMI Data: Warehouse HMI_networkHealth_pnioDevices{46}" : Push Button Data = PLC "HMI Data: Warehouse HMI".networkHealth.pnioDevices[46], 100 ms
   "HMI Data: Warehouse HMI_networkHealth_pnioDevices{47}" : Push Button Data = PLC "HMI Data: Warehouse HMI".networkHealth.pnioDevices[47], 100 ms
   "HMI Data: Warehouse HMI_networkHealth_pnioDevices{48}" : Push Button Data = PLC "HMI Data: Warehouse HMI".networkHealth.pnioDevices[48], 100 ms
   "HMI Data: Warehouse HMI_networkHealth_et200spPopUp" : Station: ET200SP Comm Debug Data = PLC "HMI Data: Warehouse HMI".networkHealth.et200spPopUp, 100 ms
   "HMI Data: Warehouse HMI_networkHealth_kp8PopUp" : Station: KP8 Comm Debug Data = PLC "HMI Data: Warehouse HMI".networkHealth.kp8PopUp, 100 ms
   "HMI Data: Warehouse HMI_networkHealth_selectedDevice" : Int = PLC "HMI Data: Warehouse HMI".networkHealth.selectedDevice, 100 ms

HMI tags "Pop Ups: Select Buttons"
   "HMI Data: Warehouse HMI_pop_up_select_buttons_buttons{0}" : Push Button Data = PLC "HMI Data: Warehouse HMI".pop_up.select_buttons.buttons[0], 100 ms
   "HMI Data: Warehouse HMI_pop_up_select_buttons_buttons{1}" : Push Button Data = PLC "HMI Data: Warehouse HMI".pop_up.select_buttons.buttons[1], 100 ms
   "HMI Data: Warehouse HMI_pop_up_select_buttons_buttons{2}" : Push Button Data = PLC "HMI Data: Warehouse HMI".pop_up.select_buttons.buttons[2], 100 ms
   "HMI Data: Warehouse HMI_pop_up_select_buttons_buttons{3}" : Push Button Data = PLC "HMI Data: Warehouse HMI".pop_up.select_buttons.buttons[3], 100 ms
   "HMI Data: Warehouse HMI_pop_up_select_buttons_buttons{4}" : Push Button Data = PLC "HMI Data: Warehouse HMI".pop_up.select_buttons.buttons[4], 100 ms
   "HMI Data: Warehouse HMI_pop_up_select_buttons_buttons{5}" : Push Button Data = PLC "HMI Data: Warehouse HMI".pop_up.select_buttons.buttons[5], 100 ms
   "HMI Data: Warehouse HMI_pop_up_select_buttons_buttons{6}" : Push Button Data = PLC "HMI Data: Warehouse HMI".pop_up.select_buttons.buttons[6], 100 ms
   "HMI Data: Warehouse HMI_pop_up_select_buttons_buttons{7}" : Push Button Data = PLC "HMI Data: Warehouse HMI".pop_up.select_buttons.buttons[7], 100 ms
   "HMI Data: Warehouse HMI_pop_up_select_buttons_close_screen" : Push Button Data = PLC "HMI Data: Warehouse HMI".pop_up.select_buttons.close_screen, 100 ms
